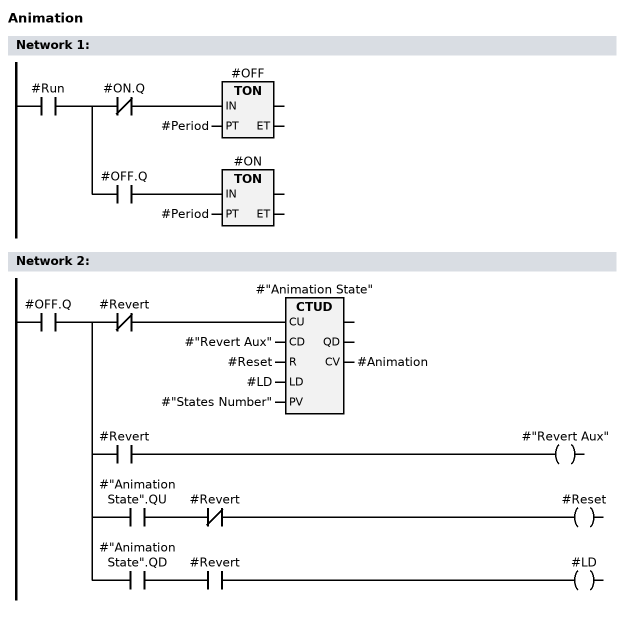
   #OFF(IN := #Run AND NOT #ON.Q, PT := #Period);   // TON
   #ON(IN := #Run AND #OFF.Q, PT := #Period);   // TON
END_REGION

REGION Network 2
   #"Animation State"(CU := #OFF.Q AND NOT #Revert,   // CTUD
                      CD := #"Revert Aux",
                      R := #Reset,
                      LD := #LD,
                      PV := #"States Number",
                      CV => #Animation);
   #"Revert Aux" := #OFF.Q AND #Revert;
   #Reset := #OFF.Q AND #"Animation State".QU AND NOT #Revert;
   #LD := #OFF.Q AND #"Animation State".QD AND #Revert;
END_REGION
END_FUNCTION_BLOCK

FUNCTION "Bool to Word" : Void   // FC202, FBD
{ S7_Optimized_Access := 'FALSE' }
VERSION : 0.1
// Die Funktion gruppiert 16 Variablen vom Datentyp "Bool" zu einer Variablen vom Datentyp "Word".
// *******************************************************************************
// The function groups 16 variables with type of data "Bool" to a variable with type of data "Word".
   VAR_INPUT
      Bit0 : Bool;
      Bit1 : Bool;
      Bit2 : Bool;
      Bit3 : Bool;
      Bit4 : Bool;
      Bit5 : Bool;
      Bit6 : Bool;
      Bit7 : Bool;
      Bit8 : Bool;
      Bit9 : Bool;
      Bit10 : Bool;
      Bit11 : Bool;
      Bit12 : Bool;
      Bit13 : Bool;
      Bit14 : Bool;
      Bit15 : Bool;
   END_VAR
   VAR_OUTPUT
      "Word" : Word;
   END_VAR
   VAR_TEMP
      aux : DInt;
   END_VAR
BEGIN

REGION Network 1: aux
   // Setze Hilfsvariable "aux" auf den Anfangswert 0.
   // ***************************************************************************
   // Set the auxiliary variable "aux" to the initial value 0.
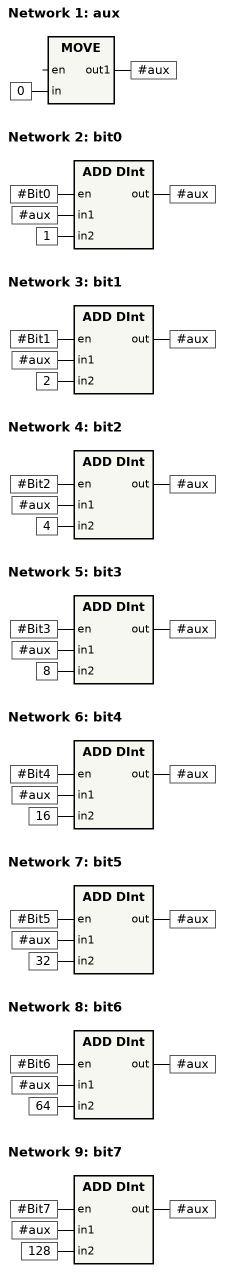
   #aux := 0;
END_REGION

REGION Network 2: bit0
   // Addiere Bit 0 zur Hilfsvariable "aux" vom Datentyp "UInt".
   // ***************************************************************************
   // Add Bit 0 to the auxiliary variable "aux" with type of data "UInt".
   IF #Bit0 THEN #aux := #aux + 1; END_IF;
END_REGION

REGION Network 3: bit1
   // Addiere Bit 1 zur Hilfsvariable "aux".
   // ***************************************************************************
   // Add Bit 1 to the auxiliary variable "aux".
   IF #Bit1 THEN #aux := #aux + 2; END_IF;
END_REGION

REGION Network 4: bit2
   // Addiere Bit 2 zur Hilfsvariable "aux".
   // ***************************************************************************
   // Add Bit 2 to the auxiliary variable "aux".
   IF #Bit2 THEN #aux := #aux + 4; END_IF;
END_REGION

REGION Network 5: bit3
   // Addiere Bit 3 zur Hilfsvariable "aux".
   // ***************************************************************************
   // Add Bit 3 to the auxiliary variable "aux".
   IF #Bit3 THEN #aux := #aux + 8; END_IF;
END_REGION

REGION Network 6: bit4
   // Addiere Bit 4 zur Hilfsvariable "aux".
   // ***************************************************************************
   // Add Bit 4 to the auxiliary variable "aux".
   IF #Bit4 THEN #aux := #aux + 16; END_IF;
END_REGION

REGION Network 7: bit5
   // Addiere Bit 5 zur Hilfsvariable "aux".
   // ***************************************************************************
   // Add Bit 5 to the auxiliary variable "aux".
   IF #Bit5 THEN #aux := #aux + 32; END_IF;
END_REGION

REGION Network 8: bit6
   // Addiere Bit 6 zur Hilfsvariable "aux".
   // ***************************************************************************
   // Add Bit 6 to the auxiliary variable "aux".
   IF #Bit6 THEN #aux := #aux + 64; END_IF;
END_REGION

REGION Network 9: bit7
   // Addiere Bit 7 zur Hilfsvariable "aux".
   // ***************************************************************************
   // Add Bit 7 to the auxiliary variable "aux".
   IF #Bit7 THEN #aux := #aux + 128; END_IF;
END_REGION

REGION Network 10: bit8
   // Addiere Bit 8 zur Hilfsvariable "aux".
   // ***************************************************************************
   // Add Bit 8 to the auxiliary variable "aux".
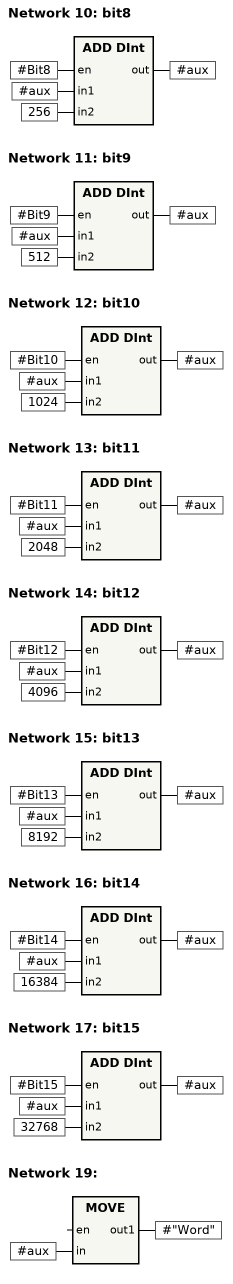
   IF #Bit8 THEN #aux := #aux + 256; END_IF;
END_REGION

REGION Network 11: bit9
   // Addiere Bit 9 zur Hilfsvariable "aux".
   // ***************************************************************************
   // Add Bit 9 to the auxiliary variable "aux".
   IF #Bit9 THEN #aux := #aux + 512; END_IF;
END_REGION

REGION Network 12: bit10
   // Addiere Bit 10 zur Hilfsvariable "aux".
   // ***************************************************************************
   // Add Bit 10 to the auxiliary variable "aux".
   IF #Bit10 THEN #aux := #aux + 1024; END_IF;
END_REGION

REGION Network 13: bit11
   // Addiere Bit 11 zur Hilfsvariable "aux".
   // ***************************************************************************
   // Add Bit 11 to the auxiliary variable "aux".
   IF #Bit11 THEN #aux := #aux + 2048; END_IF;
END_REGION

REGION Network 14: bit12
   // Addiere Bit 12 zur Hilfsvariable "aux".
   // ***************************************************************************
   // Add Bit 12 to the auxiliary variable "aux".
   IF #Bit12 THEN #aux := #aux + 4096; END_IF;
END_REGION

REGION Network 15: bit13
   // Addiere Bit 13 zur Hilfsvariable "aux".
   // ***************************************************************************
   // Add Bit 13 to the auxiliary variable "aux".
   IF #Bit13 THEN #aux := #aux + 8192; END_IF;
END_REGION

REGION Network 16: bit14
   // Addiere Bit 14 zur Hilfsvariable "aux".
   // ***************************************************************************
   // Add Bit 14 to the auxiliary variable "aux".
   IF #Bit14 THEN #aux := #aux + 16384; END_IF;
END_REGION

REGION Network 17: bit15
   // Addiere Bit 15 zur Hilfsvariable "aux".
   // ***************************************************************************
   // Add Bit 15 to the auxiliary variable "aux".
   IF #Bit15 THEN #aux := #aux + 32768; END_IF;
END_REGION

REGION Network 18: Word
   // Der Wert der Variablen "aux" wird  vom Datentyp "UInt" zum Datentyp "Word" konvertiert und der Ausgangsvariablen "Word" übergeben.
   // ***************************************************************************
   // The value of the variable "aux" will convert from type of data "UInt" to type of data "Word" and transfered to the output variable "Word".
END_REGION

REGION Network 19
   #"Word" := #aux;
END_REGION
END_FUNCTION

// folder: 60 - 69 Alarm & Status Handling

FUNCTION_BLOCK "63_E500 Fuel Pumps Not Working"   // FB63, LAD
{ S7_Optimized_Access := 'TRUE' }
VERSION : 0.1
   VAR_INPUT
      "E500A Not Runing Alarm" : Bool;
      "E500A Triped Alarm" : Bool;
      "E500B Not Runing Alarm" : Bool;
      "E500B Triped Alarm" : Bool;
      "E500A Control" : Bool;
      "E500A RUN" : Bool;
      "E500B Control" : Bool;
      "E500B RUN" : Bool;
      "Reset Alarms" : Bool;
   END_VAR
   VAR_OUTPUT
      "E500A Unavailable" : Bool;
      "E500B Unavailable" : Bool;
   END_VAR
   VAR
      IEC_Timer_0_Instance : TON_TIME;
      IEC_Timer_0_Instance_1 : TON_TIME;
      "E500A Unavailable_TP" : TP_TIME;
      "E500B Unavailable_TP" : TP_TIME;
      "E500A Unavailable Delay" : TON_TIME;
      "E500B Unavailable Delay" : TON_TIME;
      "E500A Unavailable_TOF" : TOF_TIME;
      "E500B Unavailable_TOF" : TOF_TIME;
   END_VAR
BEGIN

REGION Network 1: E500A Unavailable
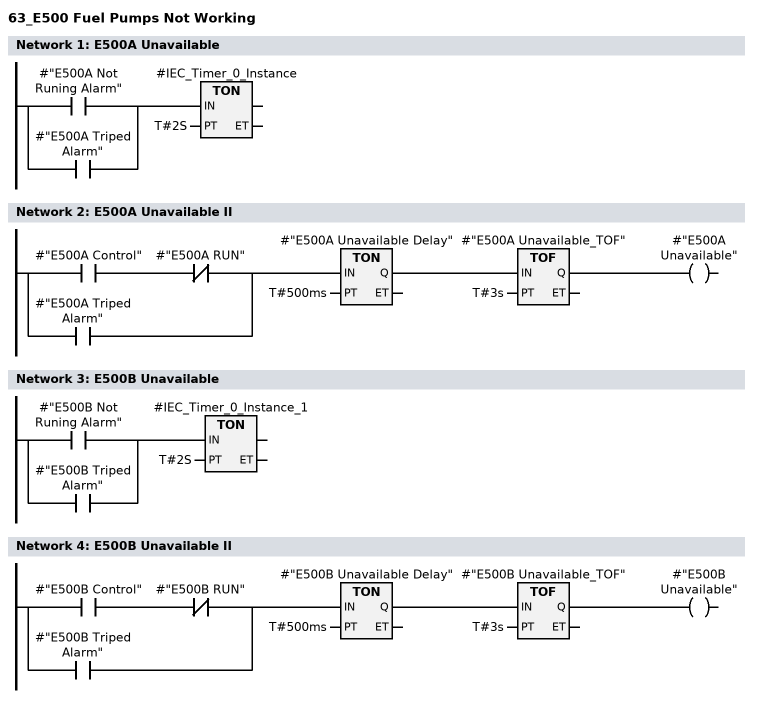
   #IEC_Timer_0_Instance(IN := #"E500A Not Runing Alarm" OR #"E500A Triped Alarm", PT := T#2S);   // TON
END_REGION

REGION Network 2: E500A Unavailable II
   #"E500A Unavailable Delay"(IN := (#"E500A Control" AND NOT #"E500A RUN") OR #"E500A Triped Alarm",   // TON
                           PT := T#500ms);
   #"E500A Unavailable_TOF"(IN := #"E500A Unavailable Delay".Q, PT := T#3s);   // TOF
   #"E500A Unavailable" := #"E500A Unavailable_TOF".Q;
END_REGION

REGION Network 3: E500B Unavailable
   #IEC_Timer_0_Instance_1(IN := #"E500B Not Runing Alarm" OR #"E500B Triped Alarm", PT := T#2S);   // TON
END_REGION

REGION Network 4: E500B Unavailable II
   #"E500B Unavailable Delay"(IN := (#"E500B Control" AND NOT #"E500B RUN") OR #"E500B Triped Alarm",   // TON
                           PT := T#500ms);
   #"E500B Unavailable_TOF"(IN := #"E500B Unavailable Delay".Q, PT := T#3s);   // TOF
   #"E500B Unavailable" := #"E500B Unavailable_TOF".Q;
END_REGION
END_FUNCTION_BLOCK

FUNCTION_BLOCK "64_Safety System Interlock"   // FB64, LAD
{ S7_Optimized_Access := 'TRUE' }
VERSION : 0.1
   VAR_INPUT
      "Safety Interlock" : Bool;
      "Reset Lockout" : Bool;
   END_VAR
   VAR_OUTPUT
      "Lockout Healthy" : Bool;
   END_VAR
   VAR
      "Interlock Fail" : Bool;
      "Aux_Interlock Fail" : Bool;
      "Initial Puls" : Bool;
      "Aux Initial Puls" : Bool;
      True : Bool;
      False : Bool;
   END_VAR
BEGIN

REGION Network 1: True/False
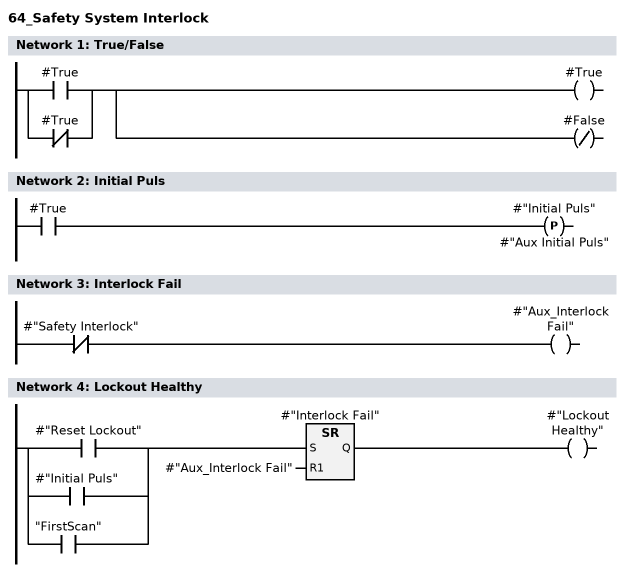
   RUNG wire#powerrail
      Contact( #True )
      wire#w1
      Coil( #True )
   END_RUNG
   RUNG wire#powerrail
      I_Contact( #True )
   END_RUNG wire#w1
   RUNG wire#w1
      I_Coil( #False )
   END_RUNG
   // the same network as SCL:
   #True := #True OR NOT #True;
   #False := NOT #True;
END_REGION

REGION Network 2: Initial Puls
   #"Initial Puls" := #True AND NOT #"Aux Initial Puls";   // rising edge
   #"Aux Initial Puls" := #True;
END_REGION

REGION Network 3: Interlock Fail
   RUNG wire#powerrail
      I_Contact( #"Safety Interlock" )
      Coil( #"Aux_Interlock Fail" )
   END_RUNG
   // the same network as SCL:
   #"Aux_Interlock Fail" := NOT #"Safety Interlock";
END_REGION

REGION Network 4: Lockout Healthy
   RUNG wire#powerrail
      Contact( #"Reset Lockout" )
      wire#w1
      S_SR(operand := #"Interlock Fail", r1 := #"Aux_Interlock Fail")
      Coil( #"Lockout Healthy" )
   END_RUNG
   RUNG wire#powerrail
      Contact( #"Initial Puls" )
   END_RUNG wire#w1
   RUNG wire#powerrail
      Contact( "FirstScan" )
   END_RUNG wire#w1
   // the same network as SCL:
   IF #"Reset Lockout" OR #"Initial Puls" OR "FirstScan" THEN
       #"Interlock Fail" := TRUE;   // SR flip-flop
   END_IF;
   IF #"Aux_Interlock Fail" THEN #"Interlock Fail" := FALSE; END_IF;
   #"Lockout Healthy" := #"Interlock Fail";
END_REGION
END_FUNCTION_BLOCK

FUNCTION "60_Alarms" : Void   // FC60, LAD
TITLE = Alarm Processing
{ S7_Optimized_Access := 'TRUE' }
AUTHOR : JRS
VERSION : 0.1
// To determine alarm conditions
   VAR_TEMP   // added for the SCL form of the ladder/FBD networks
      _w1 : Bool;
      _w2 : Bool;
      _w3 : Bool;
   END_VAR
BEGIN

REGION Network 1: DB60 DBX0.0 = Master PLC Heart Beat Missing
   // IGG_ALARM_WORD_01_BIT_0             Should be changed with the master PLC tag
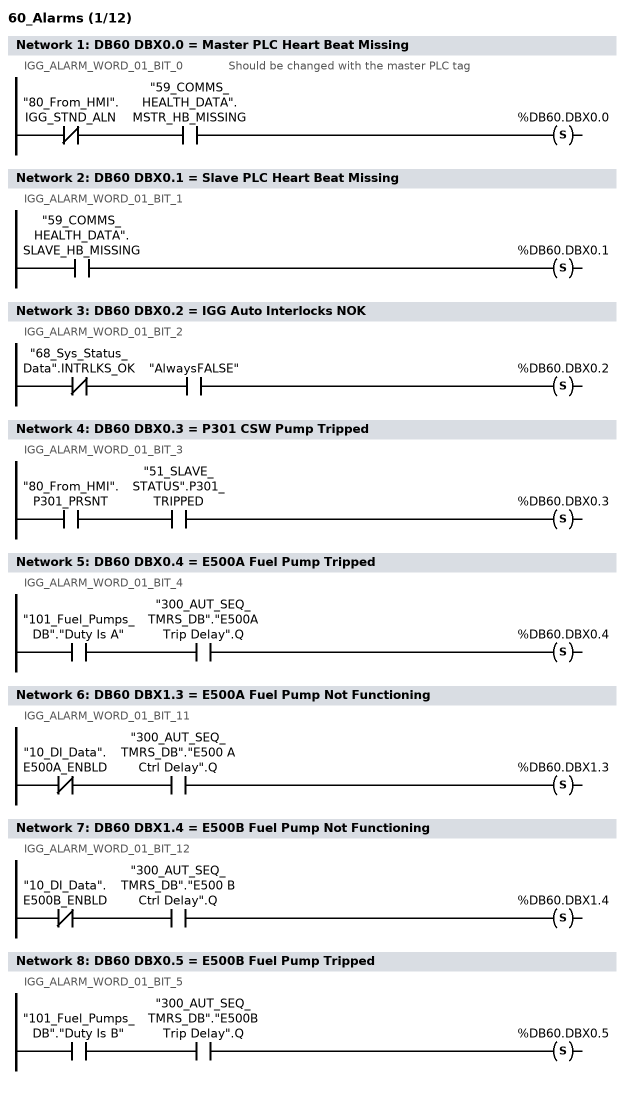
   RUNG wire#powerrail
      I_Contact( "80_From_HMI".IGG_STND_ALN )
      Contact( "59_COMMS_HEALTH_DATA".MSTR_HB_MISSING )
      S_Coil( %DB60.DBX0.0 )
   END_RUNG
   // the same network as SCL:
   IF NOT "80_From_HMI".IGG_STND_ALN AND "59_COMMS_HEALTH_DATA".MSTR_HB_MISSING THEN
       %DB60.DBX0.0 := TRUE;
   END_IF;
END_REGION

REGION Network 2: DB60 DBX0.1 = Slave PLC Heart Beat Missing
   // IGG_ALARM_WORD_01_BIT_1
   RUNG wire#powerrail
      Contact( "59_COMMS_HEALTH_DATA".SLAVE_HB_MISSING )
      S_Coil( %DB60.DBX0.1 )
   END_RUNG
   // the same network as SCL:
   IF "59_COMMS_HEALTH_DATA".SLAVE_HB_MISSING THEN %DB60.DBX0.1 := TRUE; END_IF;
END_REGION

REGION Network 3: DB60 DBX0.2 = IGG Auto Interlocks NOK
   // IGG_ALARM_WORD_01_BIT_2
   RUNG wire#powerrail
      I_Contact( "68_Sys_Status_Data".INTRLKS_OK )
      Contact( "AlwaysFALSE" )
      S_Coil( %DB60.DBX0.2 )
   END_RUNG
   // the same network as SCL:
   IF NOT "68_Sys_Status_Data".INTRLKS_OK AND "AlwaysFALSE" THEN %DB60.DBX0.2 := TRUE; END_IF;
END_REGION

REGION Network 4: DB60 DBX0.3 = P301 CSW Pump Tripped
   // IGG_ALARM_WORD_01_BIT_3
   RUNG wire#powerrail
      Contact( "80_From_HMI".P301_PRSNT )
      Contact( "51_SLAVE_STATUS".P301_TRIPPED )
      S_Coil( %DB60.DBX0.3 )
   END_RUNG
   // the same network as SCL:
   IF "80_From_HMI".P301_PRSNT AND "51_SLAVE_STATUS".P301_TRIPPED THEN %DB60.DBX0.3 := TRUE; END_IF;
END_REGION

REGION Network 5: DB60 DBX0.4 = E500A Fuel Pump Tripped
   // IGG_ALARM_WORD_01_BIT_4
   RUNG wire#powerrail
      Contact( "101_Fuel_Pumps_DB"."Duty Is A" )
      Contact( "300_AUT_SEQ_TMRS_DB"."E500A Trip Delay".Q )
      S_Coil( %DB60.DBX0.4 )
   END_RUNG
   // the same network as SCL:
   IF "101_Fuel_Pumps_DB"."Duty Is A" AND "300_AUT_SEQ_TMRS_DB"."E500A Trip Delay".Q THEN
       %DB60.DBX0.4 := TRUE;
   END_IF;
END_REGION

REGION Network 6: DB60 DBX1.3 = E500A Fuel Pump Not Functioning
   // IGG_ALARM_WORD_01_BIT_11
   RUNG wire#powerrail
      I_Contact( "10_DI_Data".E500A_ENBLD )
      Contact( "300_AUT_SEQ_TMRS_DB"."E500 A Ctrl Delay".Q )
      S_Coil( %DB60.DBX1.3 )
   END_RUNG
   // the same network as SCL:
   IF NOT "10_DI_Data".E500A_ENBLD AND "300_AUT_SEQ_TMRS_DB"."E500 A Ctrl Delay".Q THEN
       %DB60.DBX1.3 := TRUE;
   END_IF;
END_REGION

REGION Network 7: DB60 DBX1.4 = E500B Fuel Pump Not Functioning
   // IGG_ALARM_WORD_01_BIT_12
   RUNG wire#powerrail
      I_Contact( "10_DI_Data".E500B_ENBLD )
      Contact( "300_AUT_SEQ_TMRS_DB"."E500 B Ctrl Delay".Q )
      S_Coil( %DB60.DBX1.4 )
   END_RUNG
   // the same network as SCL:
   IF NOT "10_DI_Data".E500B_ENBLD AND "300_AUT_SEQ_TMRS_DB"."E500 B Ctrl Delay".Q THEN
       %DB60.DBX1.4 := TRUE;
   END_IF;
END_REGION

REGION Network 8: DB60 DBX0.5 = E500B Fuel Pump Tripped
   // IGG_ALARM_WORD_01_BIT_5
   RUNG wire#powerrail
      Contact( "101_Fuel_Pumps_DB"."Duty Is B" )
      Contact( "300_AUT_SEQ_TMRS_DB"."E500B Trip Delay".Q )
      S_Coil( %DB60.DBX0.5 )
   END_RUNG
   // the same network as SCL:
   IF "101_Fuel_Pumps_DB"."Duty Is B" AND "300_AUT_SEQ_TMRS_DB"."E500B Trip Delay".Q THEN
       %DB60.DBX0.5 := TRUE;
   END_IF;
END_REGION

REGION Network 9: DB60.DBX0.6 = E139 CAB Inverter Fault
   // IGG_ALARM_WORD_01_BIT_6
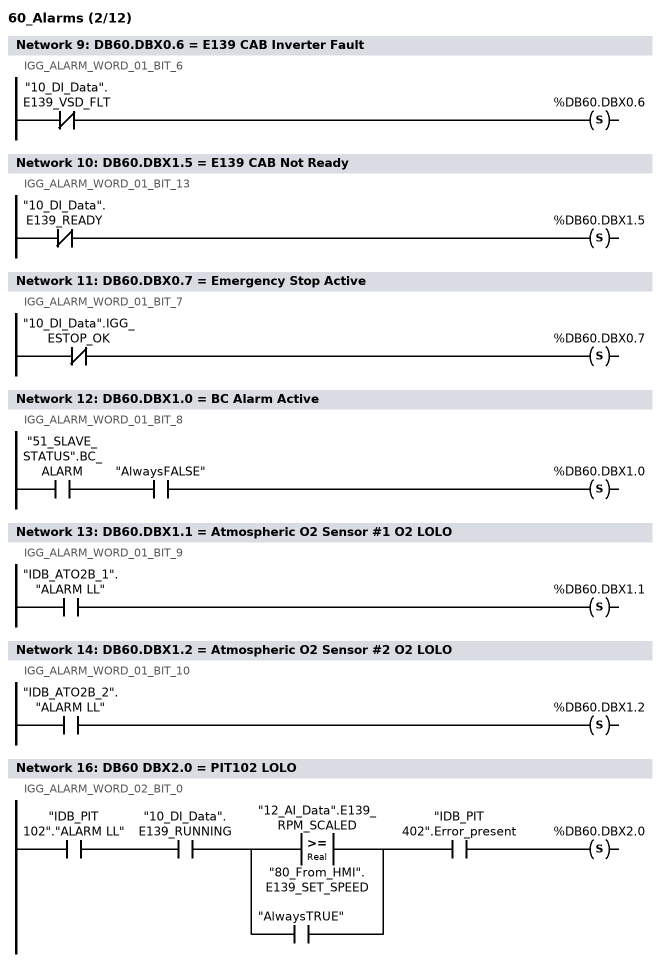
   RUNG wire#powerrail
      I_Contact( "10_DI_Data".E139_VSD_FLT )
      S_Coil( %DB60.DBX0.6 )
   END_RUNG
   // the same network as SCL:
   IF NOT "10_DI_Data".E139_VSD_FLT THEN %DB60.DBX0.6 := TRUE; END_IF;
END_REGION

REGION Network 10: DB60.DBX1.5 = E139 CAB Not Ready
   // IGG_ALARM_WORD_01_BIT_13
   RUNG wire#powerrail
      I_Contact( "10_DI_Data".E139_READY )
      S_Coil( %DB60.DBX1.5 )
   END_RUNG
   // the same network as SCL:
   IF NOT "10_DI_Data".E139_READY THEN %DB60.DBX1.5 := TRUE; END_IF;
END_REGION

REGION Network 11: DB60.DBX0.7 = Emergency Stop Active
   // IGG_ALARM_WORD_01_BIT_7
   RUNG wire#powerrail
      I_Contact( "10_DI_Data".IGG_ESTOP_OK )
      S_Coil( %DB60.DBX0.7 )
   END_RUNG
   // the same network as SCL:
   IF NOT "10_DI_Data".IGG_ESTOP_OK THEN %DB60.DBX0.7 := TRUE; END_IF;
END_REGION

REGION Network 12: DB60.DBX1.0 = BC Alarm Active
   // IGG_ALARM_WORD_01_BIT_8
   RUNG wire#powerrail
      Contact( "51_SLAVE_STATUS".BC_ALARM )
      Contact( "AlwaysFALSE" )
      S_Coil( %DB60.DBX1.0 )
   END_RUNG
   // the same network as SCL:
   IF "51_SLAVE_STATUS".BC_ALARM AND "AlwaysFALSE" THEN %DB60.DBX1.0 := TRUE; END_IF;
END_REGION

REGION Network 13: DB60.DBX1.1 = Atmospheric O2 Sensor #1 O2 LOLO
   // IGG_ALARM_WORD_01_BIT_9
   RUNG wire#powerrail
      Contact( "IDB_ATO2B_1"."ALARM LL" )
      S_Coil( %DB60.DBX1.1 )
   END_RUNG
   // the same network as SCL:
   IF "IDB_ATO2B_1"."ALARM LL" THEN %DB60.DBX1.1 := TRUE; END_IF;
END_REGION

REGION Network 14: DB60.DBX1.2 = Atmospheric O2 Sensor #2 O2 LOLO
   // IGG_ALARM_WORD_01_BIT_10
   RUNG wire#powerrail
      Contact( "IDB_ATO2B_2"."ALARM LL" )
      S_Coil( %DB60.DBX1.2 )
   END_RUNG
   // the same network as SCL:
   IF "IDB_ATO2B_2"."ALARM LL" THEN %DB60.DBX1.2 := TRUE; END_IF;
END_REGION

REGION Network 16: DB60 DBX2.0 = PIT102 LOLO
   // IGG_ALARM_WORD_02_BIT_0
   RUNG wire#powerrail
      Contact( "IDB_PIT 102"."ALARM LL" )
      Contact( "10_DI_Data".E139_RUNNING )
      wire#w1
      { S7_Templates := "SrcType := Real" } GE_Contact(in1 := "12_AI_Data".E139_RPM_SCALED, in2 := "80_From_HMI".E139_SET_SPEED)
      wire#w2
      Contact( "IDB_PIT 402".Error_present )
      S_Coil( %DB60.DBX2.0 )
   END_RUNG
   RUNG wire#w1
      Contact( "AlwaysTRUE" )
   END_RUNG wire#w2
   // the same network as SCL:
   IF "IDB_PIT 102"."ALARM LL" AND "10_DI_Data".E139_RUNNING AND (("12_AI_Data".E139_RPM_SCALED >= "80_From_HMI".E139_SET_SPEED) OR "AlwaysTRUE") AND "IDB_PIT 402".Error_present THEN
       %DB60.DBX2.0 := TRUE;
   END_IF;
END_REGION

REGION Network 17: DB60 DBX2.1 = PIT102 FAULT CA Pressure
   // IGG_ALARM_WORD_02_BIT_1
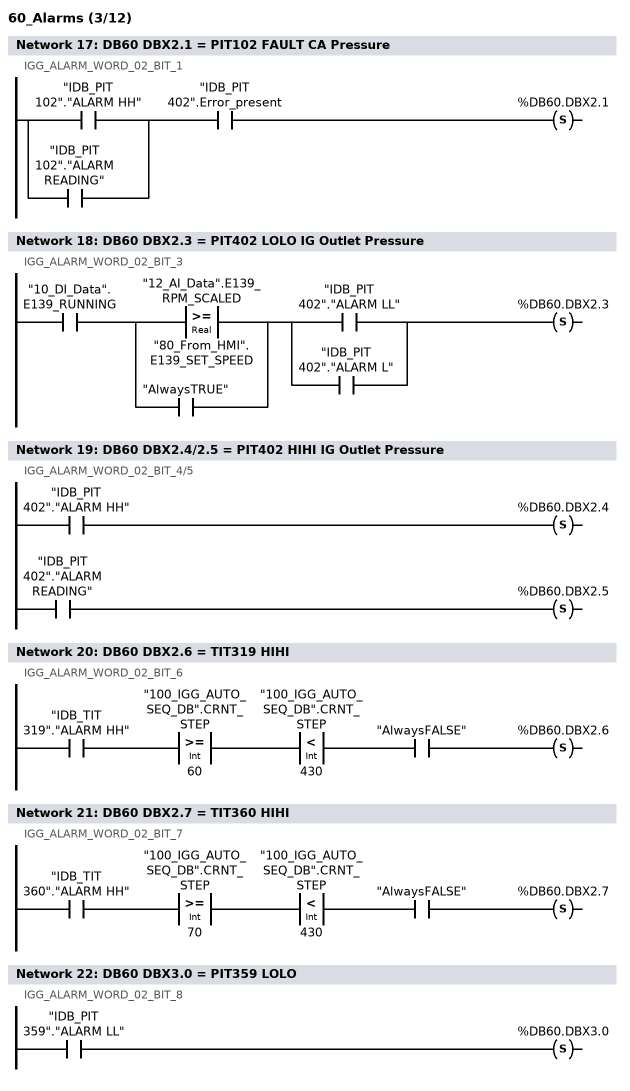
   RUNG wire#powerrail
      Contact( "IDB_PIT 102"."ALARM HH" )
      wire#w1
      Contact( "IDB_PIT 402".Error_present )
      S_Coil( %DB60.DBX2.1 )
   END_RUNG
   RUNG wire#powerrail
      Contact( "IDB_PIT 102"."ALARM READING" )
   END_RUNG wire#w1
   // the same network as SCL:
   IF ("IDB_PIT 102"."ALARM HH" OR "IDB_PIT 102"."ALARM READING") AND "IDB_PIT 402".Error_present THEN
       %DB60.DBX2.1 := TRUE;
   END_IF;
END_REGION

REGION Network 18: DB60 DBX2.3 = PIT402 LOLO IG Outlet Pressure
   // IGG_ALARM_WORD_02_BIT_3
   RUNG wire#powerrail
      Contact( "10_DI_Data".E139_RUNNING )
      wire#w1
      { S7_Templates := "SrcType := Real" } GE_Contact(in1 := "12_AI_Data".E139_RPM_SCALED, in2 := "80_From_HMI".E139_SET_SPEED)
      wire#w2
      Contact( "IDB_PIT 402"."ALARM LL" )
      wire#w3
      S_Coil( %DB60.DBX2.3 )
   END_RUNG
   RUNG wire#w1
      Contact( "AlwaysTRUE" )
   END_RUNG wire#w2
   RUNG wire#w2
      Contact( "IDB_PIT 402"."ALARM L" )
   END_RUNG wire#w3
   // the same network as SCL:
   IF "10_DI_Data".E139_RUNNING AND (("12_AI_Data".E139_RPM_SCALED >= "80_From_HMI".E139_SET_SPEED) OR "AlwaysTRUE") AND ("IDB_PIT 402"."ALARM LL" OR "IDB_PIT 402"."ALARM L") THEN
       %DB60.DBX2.3 := TRUE;
   END_IF;
END_REGION

REGION Network 19: DB60 DBX2.4/2.5 = PIT402 HIHI IG Outlet Pressure
   // IGG_ALARM_WORD_02_BIT_4/5
   RUNG wire#powerrail
      Contact( "IDB_PIT 402"."ALARM HH" )
      S_Coil( %DB60.DBX2.4 )
   END_RUNG
   RUNG wire#powerrail
      Contact( "IDB_PIT 402"."ALARM READING" )
      S_Coil( %DB60.DBX2.5 )
   END_RUNG
   // the same network as SCL:
   IF "IDB_PIT 402"."ALARM HH" THEN %DB60.DBX2.4 := TRUE; END_IF;
   IF "IDB_PIT 402"."ALARM READING" THEN %DB60.DBX2.5 := TRUE; END_IF;
END_REGION

REGION Network 20: DB60 DBX2.6 = TIT319 HIHI
   // IGG_ALARM_WORD_02_BIT_6
   RUNG wire#powerrail
      Contact( "IDB_TIT 319"."ALARM HH" )
      { S7_Templates := "SrcType := Int" } GE_Contact(in1 := "100_IGG_AUTO_SEQ_DB".CRNT_STEP, in2 := 60)
      { S7_Templates := "SrcType := Int" } LT_Contact(in1 := "100_IGG_AUTO_SEQ_DB".CRNT_STEP, in2 := 430)
      Contact( "AlwaysFALSE" )
      S_Coil( %DB60.DBX2.6 )
   END_RUNG
   // the same network as SCL:
   IF "IDB_TIT 319"."ALARM HH" AND ("100_IGG_AUTO_SEQ_DB".CRNT_STEP >= 60) AND ("100_IGG_AUTO_SEQ_DB".CRNT_STEP < 430) AND "AlwaysFALSE" THEN
       %DB60.DBX2.6 := TRUE;
   END_IF;
END_REGION

REGION Network 21: DB60 DBX2.7 = TIT360 HIHI
   // IGG_ALARM_WORD_02_BIT_7
   RUNG wire#powerrail
      Contact( "IDB_TIT 360"."ALARM HH" )
      { S7_Templates := "SrcType := Int" } GE_Contact(in1 := "100_IGG_AUTO_SEQ_DB".CRNT_STEP, in2 := 70)
      { S7_Templates := "SrcType := Int" } LT_Contact(in1 := "100_IGG_AUTO_SEQ_DB".CRNT_STEP, in2 := 430)
      Contact( "AlwaysFALSE" )
      S_Coil( %DB60.DBX2.7 )
   END_RUNG
   // the same network as SCL:
   IF "IDB_TIT 360"."ALARM HH" AND ("100_IGG_AUTO_SEQ_DB".CRNT_STEP >= 70) AND ("100_IGG_AUTO_SEQ_DB".CRNT_STEP < 430) AND "AlwaysFALSE" THEN
       %DB60.DBX2.7 := TRUE;
   END_IF;
END_REGION

REGION Network 22: DB60 DBX3.0 = PIT359 LOLO
   // IGG_ALARM_WORD_02_BIT_8
   RUNG wire#powerrail
      Contact( "IDB_PIT 359"."ALARM LL" )
      S_Coil( %DB60.DBX3.0 )
   END_RUNG
   // the same network as SCL:
   IF "IDB_PIT 359"."ALARM LL" THEN %DB60.DBX3.0 := TRUE; END_IF;
END_REGION

REGION Network 23: DB60 DBX3.4 = PIT359 HIHI
   // IGG_ALARM_WORD_02_BIT_12
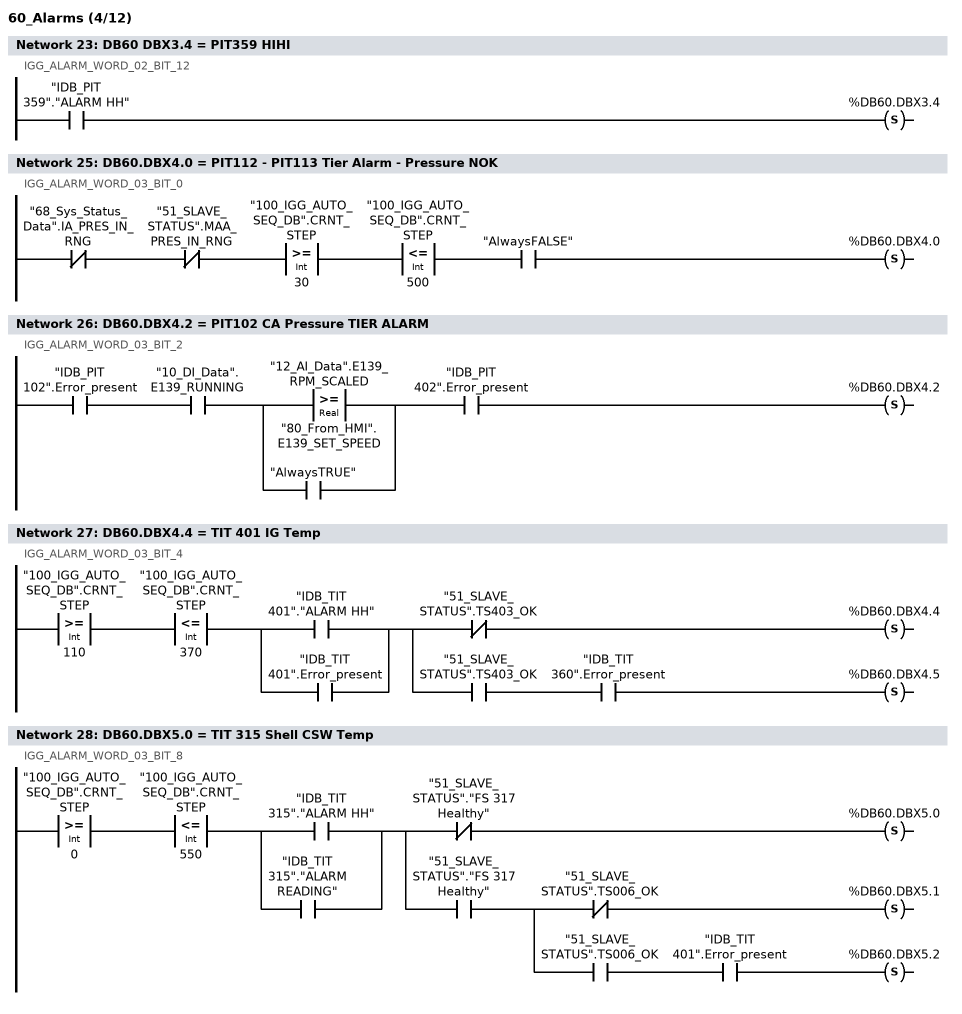
   RUNG wire#powerrail
      Contact( "IDB_PIT 359"."ALARM HH" )
      S_Coil( %DB60.DBX3.4 )
   END_RUNG
   // the same network as SCL:
   IF "IDB_PIT 359"."ALARM HH" THEN %DB60.DBX3.4 := TRUE; END_IF;
END_REGION

REGION Network 25: DB60.DBX4.0 = PIT112 - PIT113 Tier Alarm - Pressure NOK
   // IGG_ALARM_WORD_03_BIT_0
   RUNG wire#powerrail
      I_Contact( "68_Sys_Status_Data".IA_PRES_IN_RNG )
      I_Contact( "51_SLAVE_STATUS".MAA_PRES_IN_RNG )
      { S7_Templates := "SrcType := Int" } GE_Contact(in1 := "100_IGG_AUTO_SEQ_DB".CRNT_STEP, in2 := 30)
      { S7_Templates := "SrcType := Int" } LE_Contact(in1 := "100_IGG_AUTO_SEQ_DB".CRNT_STEP, in2 := 500)
      Contact( "AlwaysFALSE" )
      S_Coil( %DB60.DBX4.0 )
   END_RUNG
   // the same network as SCL:
   IF NOT "68_Sys_Status_Data".IA_PRES_IN_RNG AND NOT "51_SLAVE_STATUS".MAA_PRES_IN_RNG AND ("100_IGG_AUTO_SEQ_DB".CRNT_STEP >= 30) AND ("100_IGG_AUTO_SEQ_DB".CRNT_STEP <= 500) AND "AlwaysFALSE" THEN
       %DB60.DBX4.0 := TRUE;
   END_IF;
END_REGION

REGION Network 26: DB60.DBX4.2 = PIT102 CA Pressure TIER ALARM
   // IGG_ALARM_WORD_03_BIT_2
   RUNG wire#powerrail
      Contact( "IDB_PIT 102".Error_present )
      Contact( "10_DI_Data".E139_RUNNING )
      wire#w1
      { S7_Templates := "SrcType := Real" } GE_Contact(in1 := "12_AI_Data".E139_RPM_SCALED, in2 := "80_From_HMI".E139_SET_SPEED)
      wire#w2
      Contact( "IDB_PIT 402".Error_present )
      S_Coil( %DB60.DBX4.2 )
   END_RUNG
   RUNG wire#w1
      Contact( "AlwaysTRUE" )
   END_RUNG wire#w2
   // the same network as SCL:
   IF "IDB_PIT 102".Error_present AND "10_DI_Data".E139_RUNNING AND (("12_AI_Data".E139_RPM_SCALED >= "80_From_HMI".E139_SET_SPEED) OR "AlwaysTRUE") AND "IDB_PIT 402".Error_present THEN
       %DB60.DBX4.2 := TRUE;
   END_IF;
END_REGION

REGION Network 27: DB60.DBX4.4 = TIT 401 IG Temp
   // IGG_ALARM_WORD_03_BIT_4
   RUNG wire#powerrail
      { S7_Templates := "SrcType := Int" } GE_Contact(in1 := "100_IGG_AUTO_SEQ_DB".CRNT_STEP, in2 := 110)
      { S7_Templates := "SrcType := Int" } LE_Contact(in1 := "100_IGG_AUTO_SEQ_DB".CRNT_STEP, in2 := 370)
      wire#w1
      Contact( "IDB_TIT 401"."ALARM HH" )
      wire#w2
      I_Contact( "51_SLAVE_STATUS".TS403_OK )
      S_Coil( %DB60.DBX4.4 )
   END_RUNG
   RUNG wire#w1
      Contact( "IDB_TIT 401".Error_present )
   END_RUNG wire#w2
   RUNG wire#w2
      Contact( "51_SLAVE_STATUS".TS403_OK )
      Contact( "IDB_TIT 360".Error_present )
      S_Coil( %DB60.DBX4.5 )
   END_RUNG
   // the same network as SCL:
   #_w1 := ("100_IGG_AUTO_SEQ_DB".CRNT_STEP >= 110) AND ("100_IGG_AUTO_SEQ_DB".CRNT_STEP <= 370) AND ("IDB_TIT 401"."ALARM HH" OR "IDB_TIT 401".Error_present);
   IF #_w1 AND NOT "51_SLAVE_STATUS".TS403_OK THEN %DB60.DBX4.4 := TRUE; END_IF;
   IF #_w1 AND "51_SLAVE_STATUS".TS403_OK AND "IDB_TIT 360".Error_present THEN %DB60.DBX4.5 := TRUE; END_IF;
END_REGION

REGION Network 28: DB60.DBX5.0 = TIT 315 Shell CSW Temp
   // IGG_ALARM_WORD_03_BIT_8
   RUNG wire#powerrail
      { S7_Templates := "SrcType := Int" } GE_Contact(in1 := "100_IGG_AUTO_SEQ_DB".CRNT_STEP, in2 := 0)
      { S7_Templates := "SrcType := Int" } LE_Contact(in1 := "100_IGG_AUTO_SEQ_DB".CRNT_STEP, in2 := 550)
      wire#w1
      Contact( "IDB_TIT 315"."ALARM HH" )
      wire#w2
      I_Contact( "51_SLAVE_STATUS"."FS 317 Healthy" )
      S_Coil( %DB60.DBX5.0 )
   END_RUNG
   RUNG wire#w1
      Contact( "IDB_TIT 315"."ALARM READING" )
   END_RUNG wire#w2
   RUNG wire#w2
      Contact( "51_SLAVE_STATUS"."FS 317 Healthy" )
      wire#w3
      I_Contact( "51_SLAVE_STATUS".TS006_OK )
      S_Coil( %DB60.DBX5.1 )
   END_RUNG
   RUNG wire#w3
      Contact( "51_SLAVE_STATUS".TS006_OK )
      Contact( "IDB_TIT 401".Error_present )
      S_Coil( %DB60.DBX5.2 )
   END_RUNG
   // the same network as SCL:
   #_w1 := ("100_IGG_AUTO_SEQ_DB".CRNT_STEP >= 0) AND ("100_IGG_AUTO_SEQ_DB".CRNT_STEP <= 550) AND ("IDB_TIT 315"."ALARM HH" OR "IDB_TIT 315"."ALARM READING");
   IF #_w1 AND NOT "51_SLAVE_STATUS"."FS 317 Healthy" THEN %DB60.DBX5.0 := TRUE; END_IF;
   #_w2 := #_w1 AND "51_SLAVE_STATUS"."FS 317 Healthy";
   IF #_w2 AND NOT "51_SLAVE_STATUS".TS006_OK THEN %DB60.DBX5.1 := TRUE; END_IF;
   IF #_w2 AND "51_SLAVE_STATUS".TS006_OK AND "IDB_TIT 401".Error_present THEN %DB60.DBX5.2 := TRUE; END_IF;
END_REGION

REGION Network 29: DB60.DBX5.3 = PIT 316 Outlet CSW Pressure
   // IGG_ALARM_WORD_03_BIT_11
